   YP_T21 : TIMER[30] := ([0].PRE := 1000, [1].PRE := 10000000, [2].PRE := 10000000, [3].PRE := 3000, [3].ACC := 1845, [3].EN := 1, [3].TT := 1);
   YP_T4 : TIMER[16] := ([0].PRE := 3000, [0].ACC := 368, [0].EN := 1, [0].TT := 1, [1].PRE := 10000, [2].PRE := 10000, [2].ACC := 10001, [2].EN := 1, [2].DN := 1, [3].PRE := 60000, [3].ACC := 30907, [3].EN := 1, [3].TT := 1, [4].PRE := 5000, [4].ACC := 5000, [4].EN := 1, [4].DN := 1, [5].PRE := 5000, [6].PRE := 5000, [6].ACC := 5000, [6].EN := 1, [6].DN := 1, [7].PRE := 5000, [10].PRE := 1000);   // TIMER
        [4]   // YST1 HIGH LEVEL DE-B TIMER OFF =WET
        [5]   // YST1 HIGH LEVEL DE-B TIMER
   YP_TANK_NUMBER : ALIAS FOR YP_N10[11];
   YP_TIMER_SELECTED : ALIAS FOR YP_N55[41];   // Blunger Drain Timer Select
   YP_WATER_FILL_IDLE : ALIAS FOR YP_N40[2].0;   // BLUNGER WATER FILL IDLE
   YP_WATER_FILL_RUNNING : ALIAS FOR YP_N40[2].1;   // Blunger Water Feed Running
   YP_WD : PlantItem;   // WD
   YP_WD_RawOutput : ALIAS FOR RIO_Rack_3:3:O.Data.14;   // YP_WD
   YP_YST1_ALARM : ALIAS FOR YP_N10[1].0;
   YP_YST1_HIGH_MESSAGE : ALIAS FOR YP_B92[1].0;
   YP_YST1_HL : PlantItem;   // YST1_HL
   YP_YST1_HL_ALARM : ALIAS FOR YP_N7[38].0;
   YP_YST1_HL_FLAG : ALIAS FOR YP_N7[40].0;   // YST1 HIGH LEVEL FLAG ON=WET
   YP_YST1_HL_RawInput : ALIAS FOR RIO_Rack_3:1:I.Data.1;   // YP_YST1_HL
   YP_YST1_HL_TIMER : ALIAS FOR YP_T4[4];   // YST1 HIGH LEVEL DE-B TIMER OFF =WET
   YP_YST1_HL_TIMER2 : ALIAS FOR YP_T4[5];   // YST1 HIGH LEVEL DE-B TIMER
   YP_YST2_ALARM : ALIAS FOR YP_N10[1].1;
   YP_YST2_HIGH_LEVEL_FLAG : ALIAS FOR YP_N7[40].1;   // YST2 HIGH LEVEL FLAG ON=WET
   YP_YST2_HIGH_MESSAGE : ALIAS FOR YP_B92[1].1;
   YP_YST2_HL : PlantItem;   // YST2_HL
   YP_YST2_HL_ALARM : ALIAS FOR YP_N7[38].1;
   YP_YST2_HL_RawInput : ALIAS FOR RIO_Rack_3:1:I.Data.3;   // YP_YST2_HL
   YP_YST2_HL_TIMER : ALIAS FOR YP_T4[6];
   YP_YST2_HL_TIMER2 : ALIAS FOR YP_T4[7];
   YST_BL_PMP_ON : BOOL;   // Blunger Pump
   YST_CIP_Conns_Confirmed : BOOL := 1;
   YST_Confirm_CIP_connected : BOOL;
   YST_Confirm_Vent_connected : BOOL;
   YST_Vent_Connection_Confirmed : BOOL;
   YSVFilling_transaction_locked_timer : TIMER := (PRE := 10000);
   YSVFilling_transaction_log : DINT;
   YSVFilling_transaction_log_delay : DINT;
   YSVFilling_transaction_log_Done : DINT := -1;
   YSVFilling_transaction_log_timer : TIMER := (PRE := 10000);
END_VAR

PROGRAM _1Second   (* main routine OneSecond *)

ROUTINE OneSecond   (* ladder *)
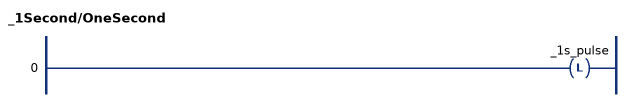
   0: OTL(_1s_pulse);
END_ROUTINE
END_PROGRAM

PROGRAM First_Task   (* main routine MainRoutine *)

ROUTINE MainRoutine   (* ladder *)
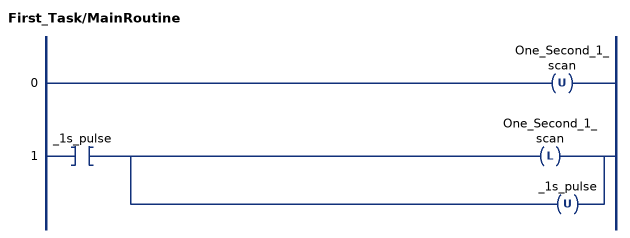
   0: OTU(One_Second_1_scan);
   1: XIC(_1s_pulse)[OTL(One_Second_1_scan) ,OTU(_1s_pulse) ];
END_ROUTINE
END_PROGRAM

PROGRAM FR_Common   (* main routine MainRoutine *)
VAR
   FR_FV31_AV08_O1 : ALIAS FOR RIO_Rack_2:12:I.Data.26;
   FR_FVS_P01_Cond_Met : BOOL;
END_VAR

ROUTINE A_FactoryTalk_Requirements   (* ladder *)
END_ROUTINE

ROUTINE Analog_scale_ftof   (* ladder *)
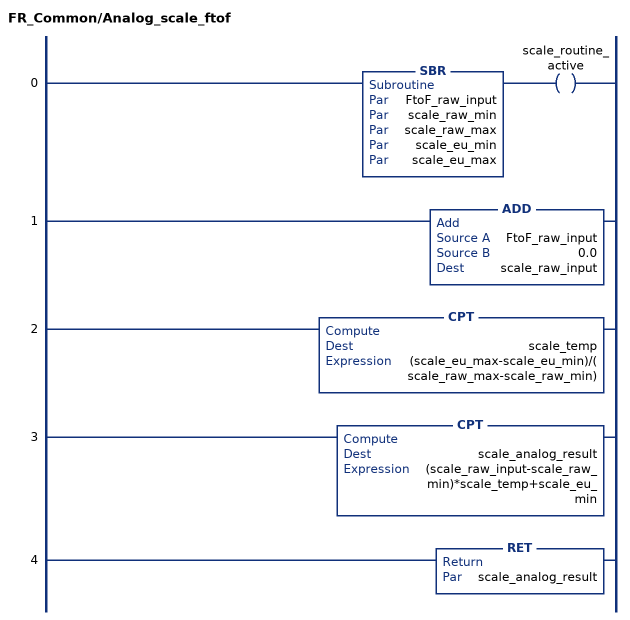
   0: SBR(FtoF_raw_input,scale_raw_min,scale_raw_max,scale_eu_min,scale_eu_max)OTE(scale_routine_active);
   1: ADD(FtoF_raw_input,0.0,scale_raw_input);
   2: CPT(scale_temp,(scale_eu_max-scale_eu_min)/(scale_raw_max-scale_raw_min));
   3: CPT(scale_analog_result,(scale_raw_input-scale_raw_min)*scale_temp+scale_eu_min);
   4: RET(scale_analog_result);
END_ROUTINE

ROUTINE Analog_Scale_FtoI   (* ladder *)
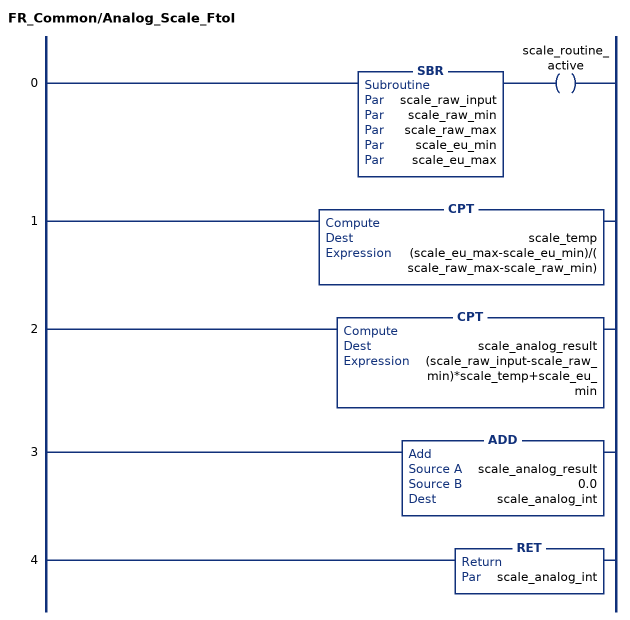
   0: SBR(scale_raw_input,scale_raw_min,scale_raw_max,scale_eu_min,scale_eu_max)OTE(scale_routine_active);
   1: CPT(scale_temp,(scale_eu_max-scale_eu_min)/(scale_raw_max-scale_raw_min));
   2: CPT(scale_analog_result,(scale_raw_input-scale_raw_min)*scale_temp+scale_eu_min);
   3: ADD(scale_analog_result,0.0,scale_analog_int);
   4: RET(scale_analog_int);
END_ROUTINE

ROUTINE Analog_Scale_ItoF   (* ladder *)
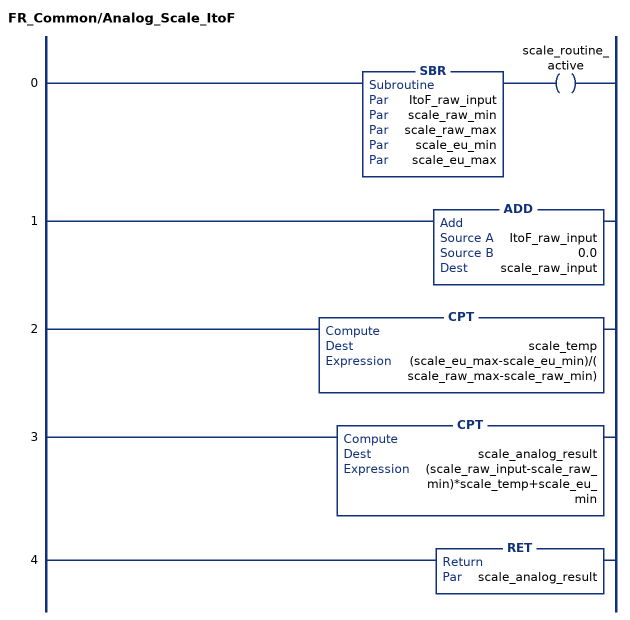
   0: SBR(ItoF_raw_input,scale_raw_min,scale_raw_max,scale_eu_min,scale_eu_max)OTE(scale_routine_active);
   1: ADD(ItoF_raw_input,0.0,scale_raw_input);
   2: CPT(scale_temp,(scale_eu_max-scale_eu_min)/(scale_raw_max-scale_raw_min));
   3: CPT(scale_analog_result,(scale_raw_input-scale_raw_min)*scale_temp+scale_eu_min);
   4: RET(scale_analog_result);
END_ROUTINE

ROUTINE Analog_Scale_ItoF_Int_Parms   (* ladder *)
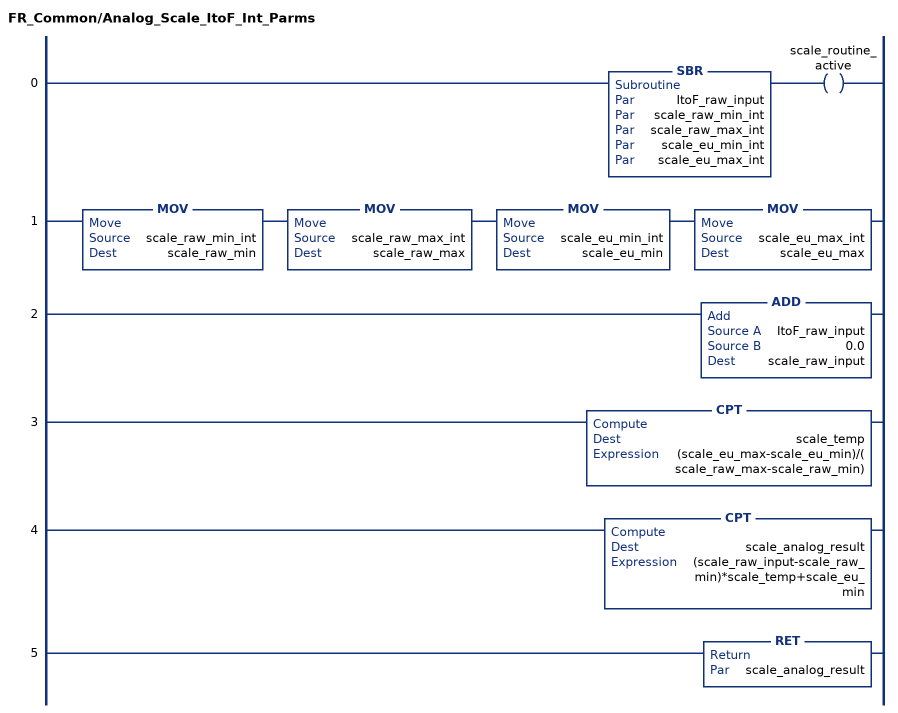
   0: SBR(ItoF_raw_input,scale_raw_min_int,scale_raw_max_int,scale_eu_min_int,scale_eu_max_int)OTE(scale_routine_active);
   1: MOV(scale_raw_min_int,scale_raw_min)MOV(scale_raw_max_int,scale_raw_max)MOV(scale_eu_min_int,scale_eu_min)MOV(scale_eu_max_int,scale_eu_max);
   2: ADD(ItoF_raw_input,0.0,scale_raw_input);
   3: CPT(scale_temp,(scale_eu_max-scale_eu_min)/(scale_raw_max-scale_raw_min));
   4: CPT(scale_analog_result,(scale_raw_input-scale_raw_min)*scale_temp+scale_eu_min);
   5: RET(scale_analog_result);
END_ROUTINE

ROUTINE FR_A_Alarms_From_PLC   (* ladder *)
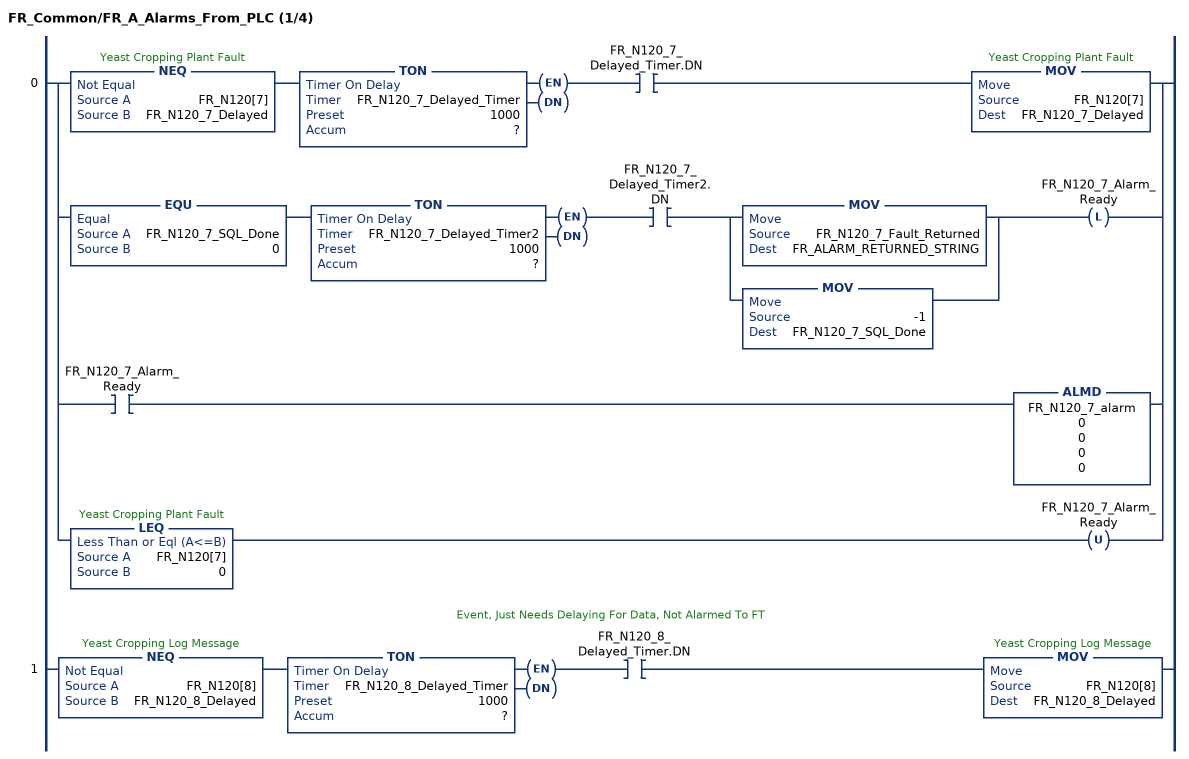
   0: [NEQ(FR_N120[7],FR_N120_7_Delayed) TON(FR_N120_7_Delayed_Timer,?,?) XIC(FR_N120_7_Delayed_Timer.DN) MOV(FR_N120[7],FR_N120_7_Delayed) ,EQU(FR_N120_7_SQL_Done,0) TON(FR_N120_7_Delayed_Timer2,?,?) XIC(FR_N120_7_Delayed_Timer2.DN) [MOV(FR_N120_7_Fault_Returned,FR_ALARM_RETURNED_STRING) ,MOV(-1,FR_N120_7_SQL_Done) ] OTL(FR_N120_7_Alarm_Ready) ,XIC(FR_N120_7_Alarm_Ready) ALMD(FR_N120_7_alarm,0,0,0,0) ,LEQ(FR_N120[7],0) OTU(FR_N120_7_Alarm_Ready) ];
   // Event, Just Needs Delaying For Data, Not Alarmed To FT
   1: NEQ(FR_N120[8],FR_N120_8_Delayed)TON(FR_N120_8_Delayed_Timer,?,?)XIC(FR_N120_8_Delayed_Timer.DN)MOV(FR_N120[8],FR_N120_8_Delayed);
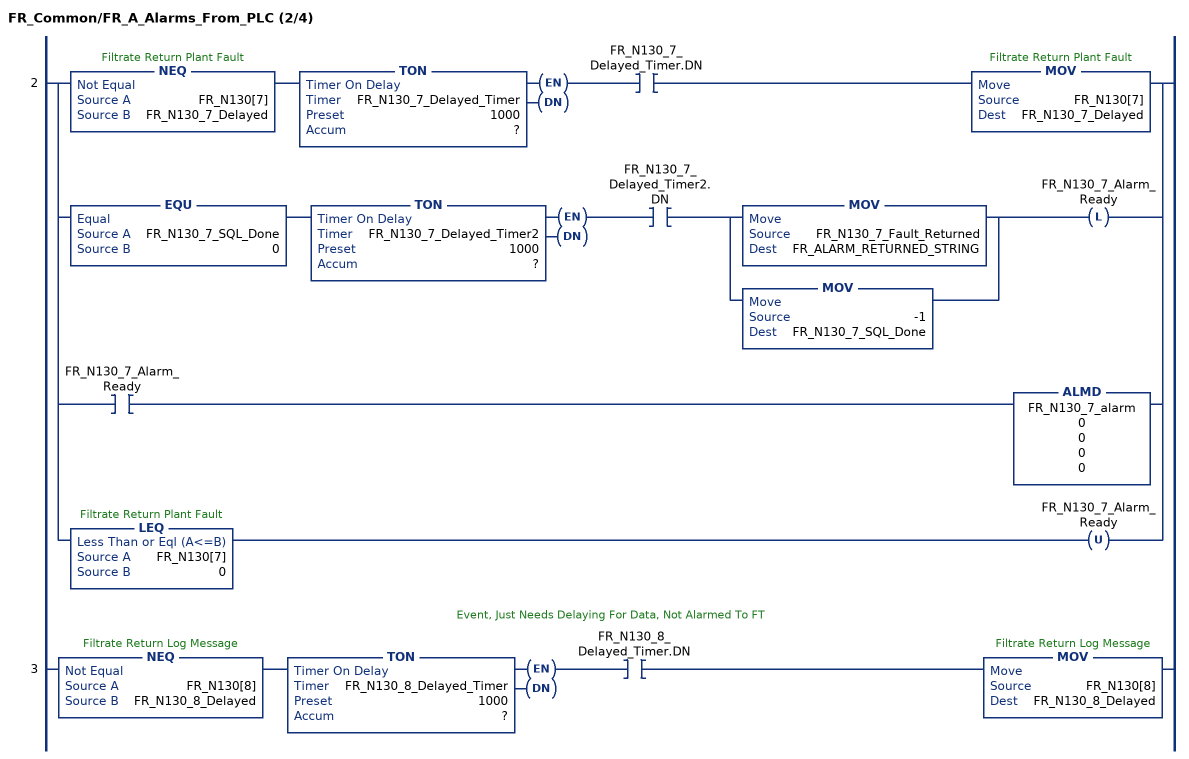
   2: [NEQ(FR_N130[7],FR_N130_7_Delayed) TON(FR_N130_7_Delayed_Timer,?,?) XIC(FR_N130_7_Delayed_Timer.DN) MOV(FR_N130[7],FR_N130_7_Delayed) ,EQU(FR_N130_7_SQL_Done,0) TON(FR_N130_7_Delayed_Timer2,?,?) XIC(FR_N130_7_Delayed_Timer2.DN) [MOV(FR_N130_7_Fault_Returned,FR_ALARM_RETURNED_STRING) ,MOV(-1,FR_N130_7_SQL_Done) ] OTL(FR_N130_7_Alarm_Ready) ,XIC(FR_N130_7_Alarm_Ready) ALMD(FR_N130_7_alarm,0,0,0,0) ,LEQ(FR_N130[7],0) OTU(FR_N130_7_Alarm_Ready) ];
   // Event, Just Needs Delaying For Data, Not Alarmed To FT
   3: NEQ(FR_N130[8],FR_N130_8_Delayed)TON(FR_N130_8_Delayed_Timer,?,?)XIC(FR_N130_8_Delayed_Timer.DN)MOV(FR_N130[8],FR_N130_8_Delayed);
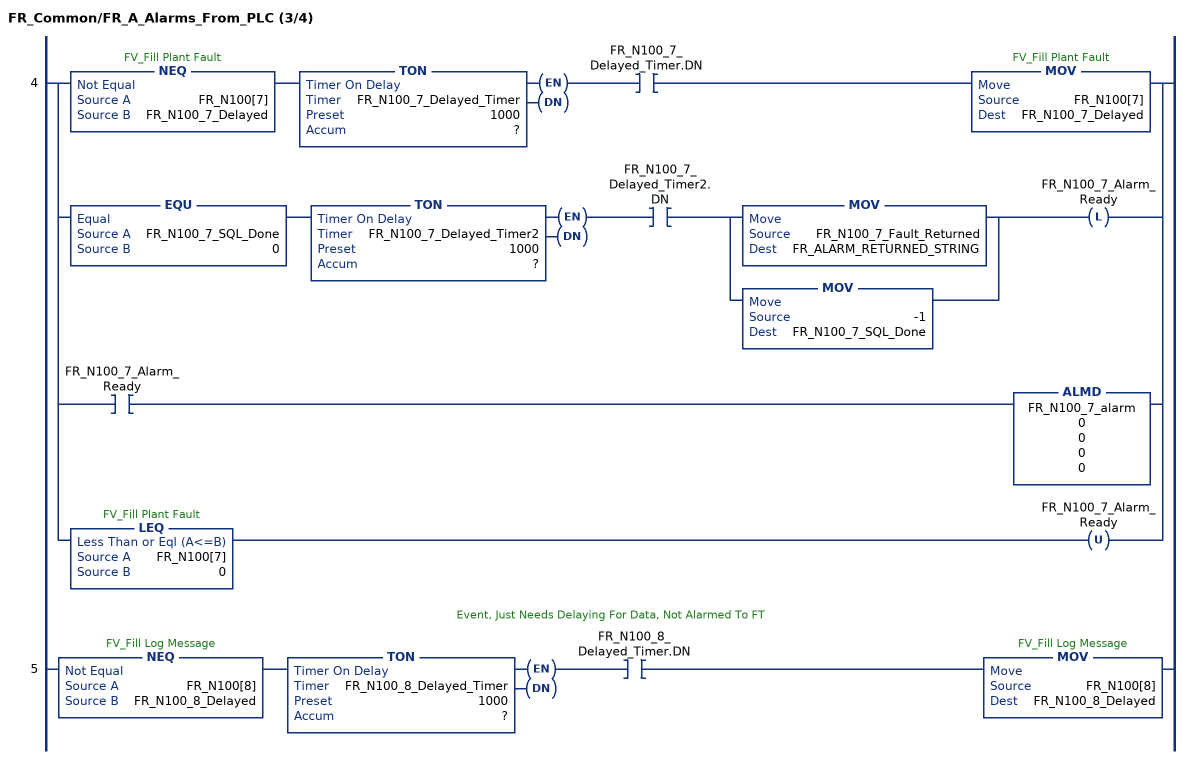
   4: [NEQ(FR_N100[7],FR_N100_7_Delayed) TON(FR_N100_7_Delayed_Timer,?,?) XIC(FR_N100_7_Delayed_Timer.DN) MOV(FR_N100[7],FR_N100_7_Delayed) ,EQU(FR_N100_7_SQL_Done,0) TON(FR_N100_7_Delayed_Timer2,?,?) XIC(FR_N100_7_Delayed_Timer2.DN) [MOV(FR_N100_7_Fault_Returned,FR_ALARM_RETURNED_STRING) ,MOV(-1,FR_N100_7_SQL_Done) ] OTL(FR_N100_7_Alarm_Ready) ,XIC(FR_N100_7_Alarm_Ready) ALMD(FR_N100_7_alarm,0,0,0,0) ,LEQ(FR_N100[7],0) OTU(FR_N100_7_Alarm_Ready) ];
   // Event, Just Needs Delaying For Data, Not Alarmed To FT
   5: NEQ(FR_N100[8],FR_N100_8_Delayed)TON(FR_N100_8_Delayed_Timer,?,?)XIC(FR_N100_8_Delayed_Timer.DN)MOV(FR_N100[8],FR_N100_8_Delayed);
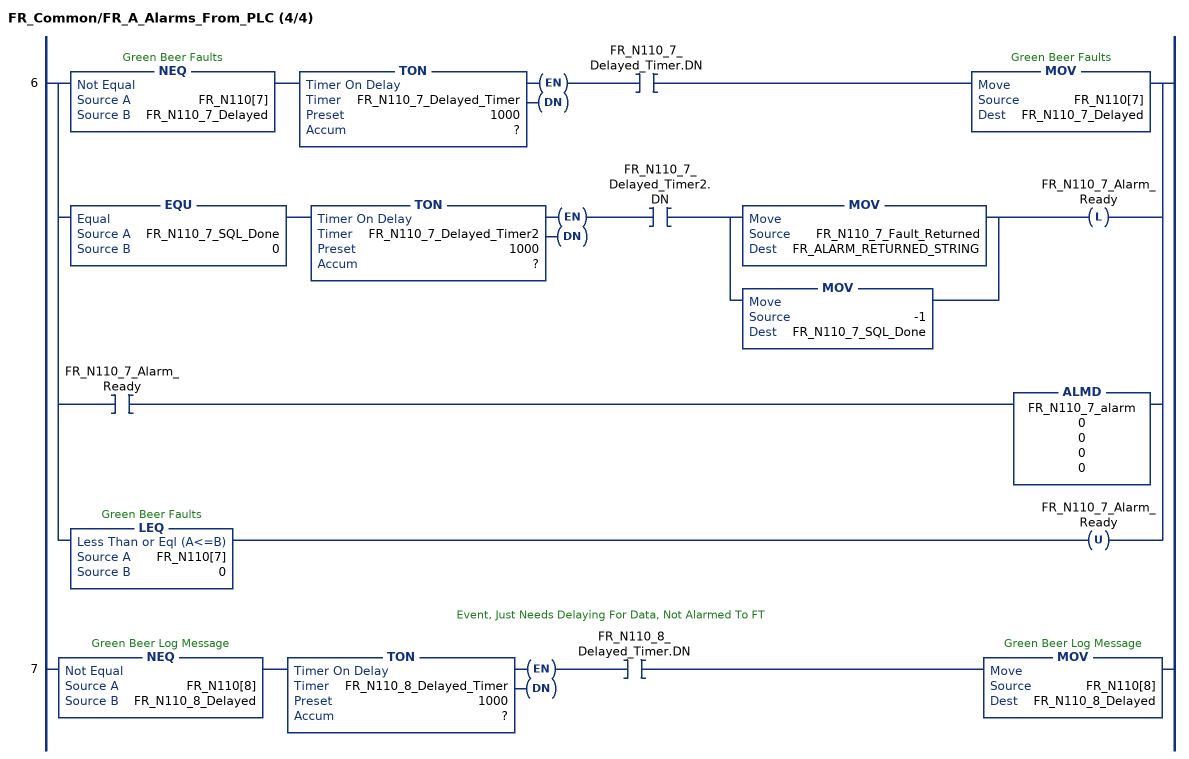
   6: [NEQ(FR_N110[7],FR_N110_7_Delayed) TON(FR_N110_7_Delayed_Timer,?,?) XIC(FR_N110_7_Delayed_Timer.DN) MOV(FR_N110[7],FR_N110_7_Delayed) ,EQU(FR_N110_7_SQL_Done,0) TON(FR_N110_7_Delayed_Timer2,?,?) XIC(FR_N110_7_Delayed_Timer2.DN) [MOV(FR_N110_7_Fault_Returned,FR_ALARM_RETURNED_STRING) ,MOV(-1,FR_N110_7_SQL_Done) ] OTL(FR_N110_7_Alarm_Ready) ,XIC(FR_N110_7_Alarm_Ready) ALMD(FR_N110_7_alarm,0,0,0,0) ,LEQ(FR_N110[7],0) OTU(FR_N110_7_Alarm_Ready) ];
   // Event, Just Needs Delaying For Data, Not Alarmed To FT
   7: NEQ(FR_N110[8],FR_N110_8_Delayed)TON(FR_N110_8_Delayed_Timer,?,?)XIC(FR_N110_8_Delayed_Timer.DN)MOV(FR_N110[8],FR_N110_8_Delayed);
END_ROUTINE

ROUTINE FR_A_Events_From_Scada   (* ladder *)
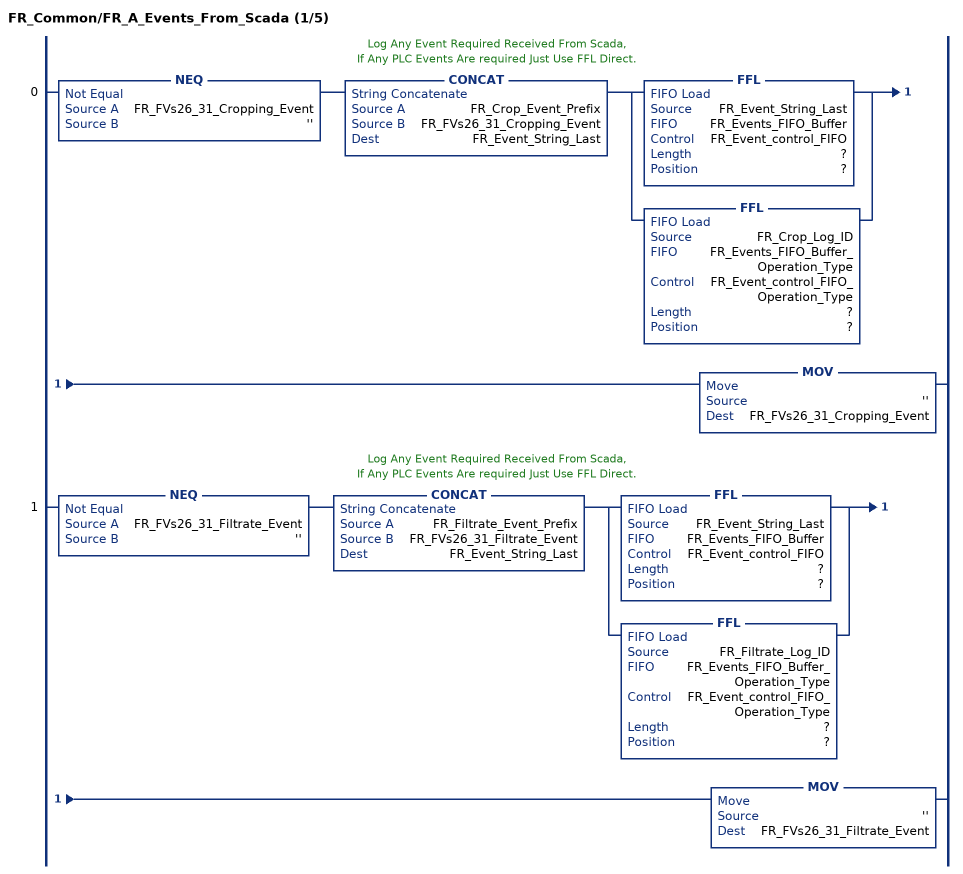
   // Log Any Event Required Received From Scada,
   // If Any PLC Events Are required Just Use FFL Direct.
   0: NEQ(FR_FVs26_31_Cropping_Event,'')CONCAT(FR_Crop_Event_Prefix,FR_FVs26_31_Cropping_Event,FR_Event_String_Last)[FFL(FR_Event_String_Last,FR_Events_FIFO_Buffer,FR_Event_control_FIFO,?,?) ,FFL(FR_Crop_Log_ID,FR_Events_FIFO_Buffer_Operation_Type,FR_Event_control_FIFO_Operation_Type,?,?) ]MOV('',FR_FVs26_31_Cropping_Event);
   // Log Any Event Required Received From Scada,
   // If Any PLC Events Are required Just Use FFL Direct.
   1: NEQ(FR_FVs26_31_Filtrate_Event,'')CONCAT(FR_Filtrate_Event_Prefix,FR_FVs26_31_Filtrate_Event,FR_Event_String_Last)[FFL(FR_Event_String_Last,FR_Events_FIFO_Buffer,FR_Event_control_FIFO,?,?) ,FFL(FR_Filtrate_Log_ID,FR_Events_FIFO_Buffer_Operation_Type,FR_Event_control_FIFO_Operation_Type,?,?) ]MOV('',FR_FVs26_31_Filtrate_Event);
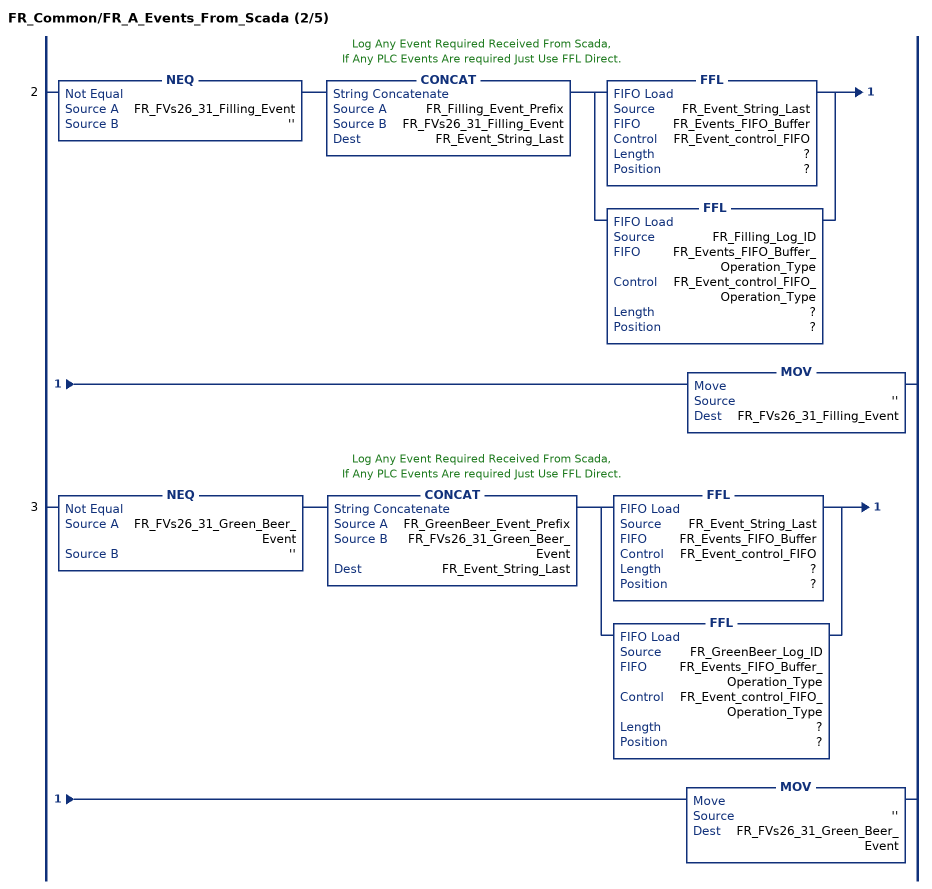
   // Log Any Event Required Received From Scada,
   // If Any PLC Events Are required Just Use FFL Direct.
   2: NEQ(FR_FVs26_31_Filling_Event,'')CONCAT(FR_Filling_Event_Prefix,FR_FVs26_31_Filling_Event,FR_Event_String_Last)[FFL(FR_Event_String_Last,FR_Events_FIFO_Buffer,FR_Event_control_FIFO,?,?) ,FFL(FR_Filling_Log_ID,FR_Events_FIFO_Buffer_Operation_Type,FR_Event_control_FIFO_Operation_Type,?,?) ]MOV('',FR_FVs26_31_Filling_Event);
   // Log Any Event Required Received From Scada,
   // If Any PLC Events Are required Just Use FFL Direct.
   3: NEQ(FR_FVs26_31_Green_Beer_Event,'')CONCAT(FR_GreenBeer_Event_Prefix,FR_FVs26_31_Green_Beer_Event,FR_Event_String_Last)[FFL(FR_Event_String_Last,FR_Events_FIFO_Buffer,FR_Event_control_FIFO,?,?) ,FFL(FR_GreenBeer_Log_ID,FR_Events_FIFO_Buffer_Operation_Type,FR_Event_control_FIFO_Operation_Type,?,?) ]MOV('',FR_FVs26_31_Green_Beer_Event);
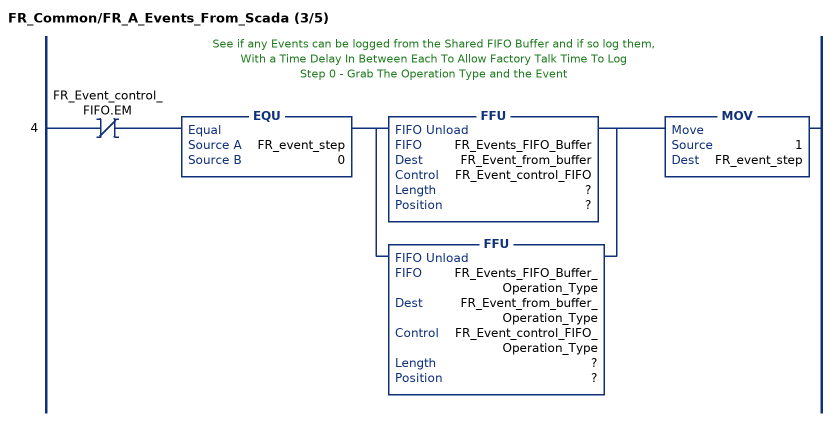
   // See if any Events can be logged from the Shared FIFO Buffer and if so log them,
   // With a Time Delay In Between Each To Allow Factory Talk Time To Log
   // Step 0 - Grab The Operation Type and the Event
   4: XIO(FR_Event_control_FIFO.EM)EQU(FR_event_step,0)[FFU(FR_Events_FIFO_Buffer,FR_Event_from_buffer,FR_Event_control_FIFO,?,?) ,FFU(FR_Events_FIFO_Buffer_Operation_Type,FR_Event_from_buffer_Operation_Type,FR_Event_control_FIFO_Operation_Type,?,?) ]MOV(1,FR_event_step);
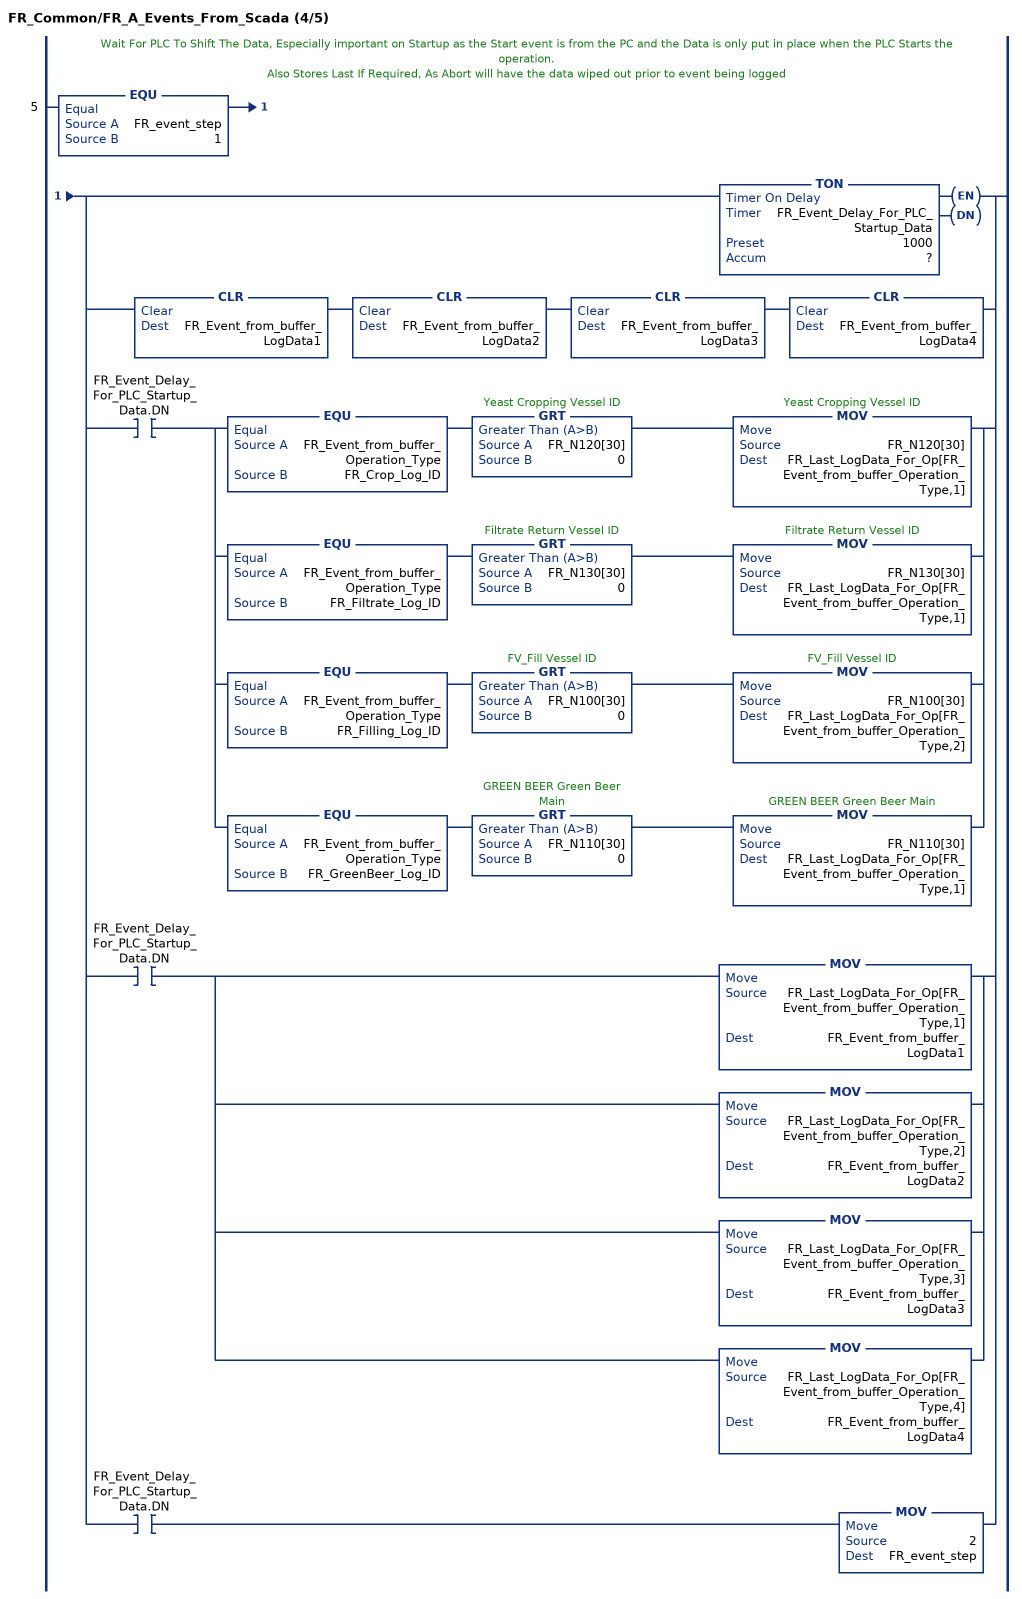
   // Wait For PLC To Shift The Data, Especially important on Startup as the Start event is from the PC and the Data is only put in place when the PLC Starts the operation.
   // Also Stores Last If Required, As Abort will have the data wiped out prior to event being logged
   5: EQU(FR_event_step,1)[TON(FR_Event_Delay_For_PLC_Startup_Data,?,?) ,CLR(FR_Event_from_buffer_LogData1) CLR(FR_Event_from_buffer_LogData2) CLR(FR_Event_from_buffer_LogData3) CLR(FR_Event_from_buffer_LogData4) ,XIC(FR_Event_Delay_For_PLC_Startup_Data.DN) [EQU(FR_Event_from_buffer_Operation_Type,FR_Crop_Log_ID) GRT(FR_N120[30],0) MOV(FR_N120[30],FR_Last_LogData_For_Op[FR_Event_from_buffer_Operation_Type,1]) ,EQU(FR_Event_from_buffer_Operation_Type,FR_Filtrate_Log_ID) GRT(FR_N130[30],0) MOV(FR_N130[30],FR_Last_LogData_For_Op[FR_Event_from_buffer_Operation_Type,1]) ,EQU(FR_Event_from_buffer_Operation_Type,FR_Filling_Log_ID) GRT(FR_N100[30],0) MOV(FR_N100[30],FR_Last_LogData_For_Op[FR_Event_from_buffer_Operation_Type,2]) ,EQU(FR_Event_from_buffer_Operation_Type,FR_GreenBeer_Log_ID) GRT(FR_N110[30],0) MOV(FR_N110[30],FR_Last_LogData_For_Op[FR_Event_from_buffer_Operation_Type,1]) ] ,XIC(FR_Event_Delay_For_PLC_Startup_Data.DN) [MOV(FR_Last_LogData_For_Op[FR_Event_from_buffer_Operation_Type,1],FR_Event_from_buffer_LogData1) ,MOV(FR_Last_LogData_For_Op[FR_Event_from_buffer_Operation_Type,2],FR_Event_from_buffer_LogData2) ,MOV(FR_Last_LogData_For_Op[FR_Event_from_buffer_Operation_Type,3],FR_Event_from_buffer_LogData3) ,MOV(FR_Last_LogData_For_Op[FR_Event_from_buffer_Operation_Type,4],FR_Event_from_buffer_LogData4) ] ,XIC(FR_Event_Delay_For_PLC_Startup_Data.DN) MOV(2,FR_event_step) ];
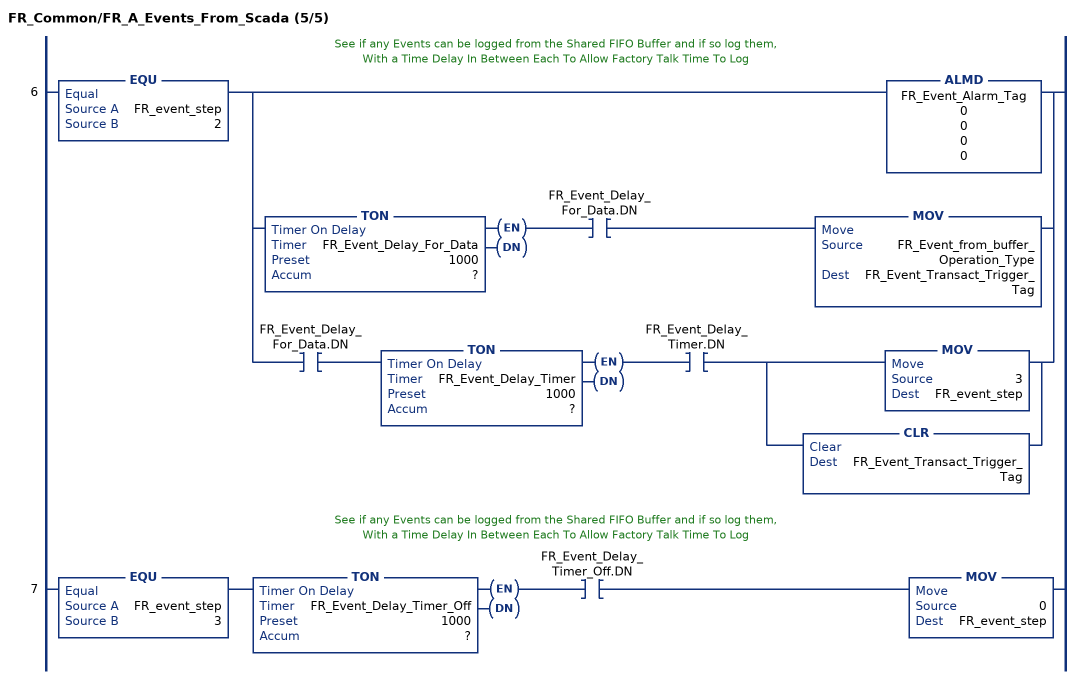
   // See if any Events can be logged from the Shared FIFO Buffer and if so log them,
   // With a Time Delay In Between Each To Allow Factory Talk Time To Log
   6: EQU(FR_event_step,2)[ALMD(FR_Event_Alarm_Tag,0,0,0,0) ,TON(FR_Event_Delay_For_Data,?,?) XIC(FR_Event_Delay_For_Data.DN) MOV(FR_Event_from_buffer_Operation_Type,FR_Event_Transact_Trigger_Tag) ,XIC(FR_Event_Delay_For_Data.DN) TON(FR_Event_Delay_Timer,?,?) XIC(FR_Event_Delay_Timer.DN) [MOV(3,FR_event_step) ,CLR(FR_Event_Transact_Trigger_Tag) ] ];
   // See if any Events can be logged from the Shared FIFO Buffer and if so log them,
   // With a Time Delay In Between Each To Allow Factory Talk Time To Log
   7: EQU(FR_event_step,3)TON(FR_Event_Delay_Timer_Off,?,?)XIC(FR_Event_Delay_Timer_Off.DN)MOV(0,FR_event_step);
END_ROUTINE

ROUTINE FR_A_Events_From_Scada_IDs   (* ladder *)
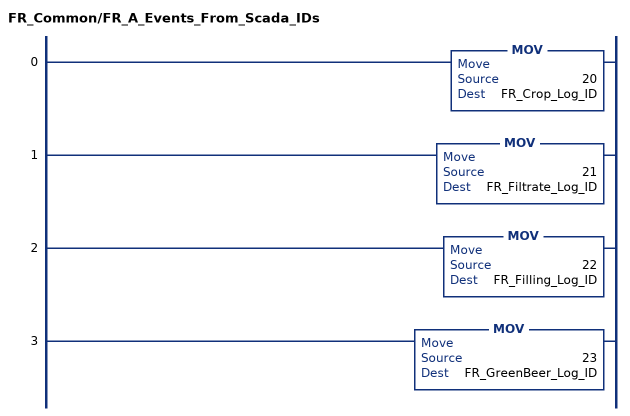
   0: MOV(20,FR_Crop_Log_ID);
   1: MOV(21,FR_Filtrate_Log_ID);
   2: MOV(22,FR_Filling_Log_ID);
   3: MOV(23,FR_GreenBeer_Log_ID);
END_ROUTINE

ROUTINE FR_A_Warnings_From_PLC   (* ladder *)
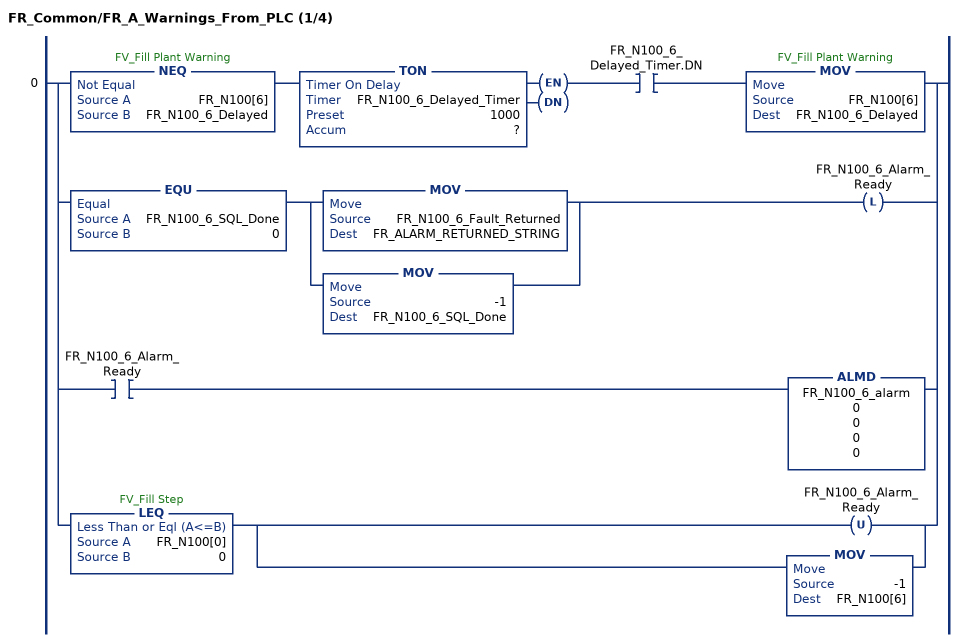
   0: [NEQ(FR_N100[6],FR_N100_6_Delayed) TON(FR_N100_6_Delayed_Timer,?,?) XIC(FR_N100_6_Delayed_Timer.DN) MOV(FR_N100[6],FR_N100_6_Delayed) ,EQU(FR_N100_6_SQL_Done,0) [MOV(FR_N100_6_Fault_Returned,FR_ALARM_RETURNED_STRING) ,MOV(-1,FR_N100_6_SQL_Done) ] OTL(FR_N100_6_Alarm_Ready) ,XIC(FR_N100_6_Alarm_Ready) ALMD(FR_N100_6_alarm,0,0,0,0) ,LEQ(FR_N100[0],0) [OTU(FR_N100_6_Alarm_Ready) ,MOV(-1,FR_N100[6]) ] ];
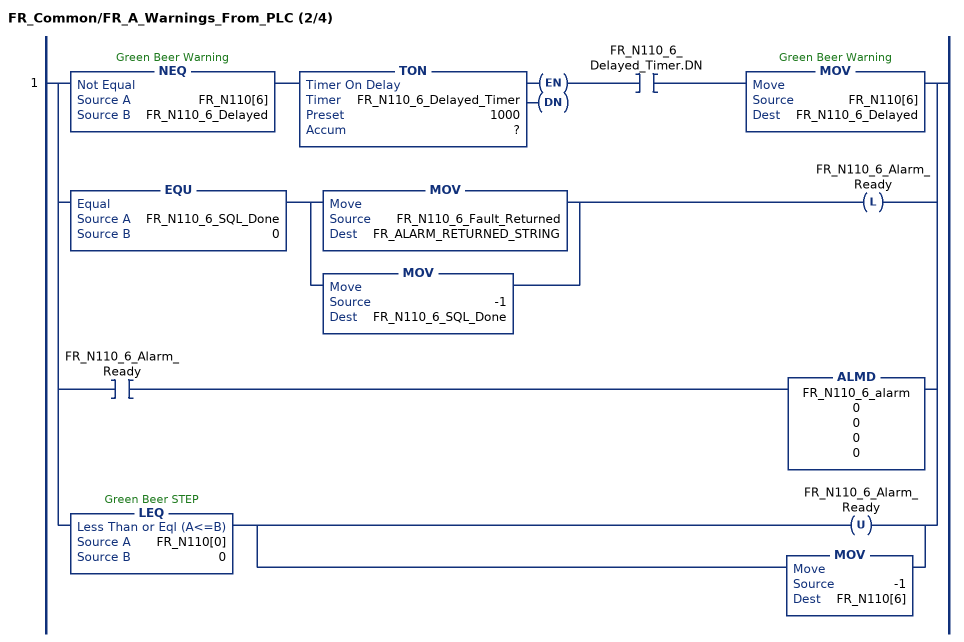
   1: [NEQ(FR_N110[6],FR_N110_6_Delayed) TON(FR_N110_6_Delayed_Timer,?,?) XIC(FR_N110_6_Delayed_Timer.DN) MOV(FR_N110[6],FR_N110_6_Delayed) ,EQU(FR_N110_6_SQL_Done,0) [MOV(FR_N110_6_Fault_Returned,FR_ALARM_RETURNED_STRING) ,MOV(-1,FR_N110_6_SQL_Done) ] OTL(FR_N110_6_Alarm_Ready) ,XIC(FR_N110_6_Alarm_Ready) ALMD(FR_N110_6_alarm,0,0,0,0) ,LEQ(FR_N110[0],0) [OTU(FR_N110_6_Alarm_Ready) ,MOV(-1,FR_N110[6]) ] ];
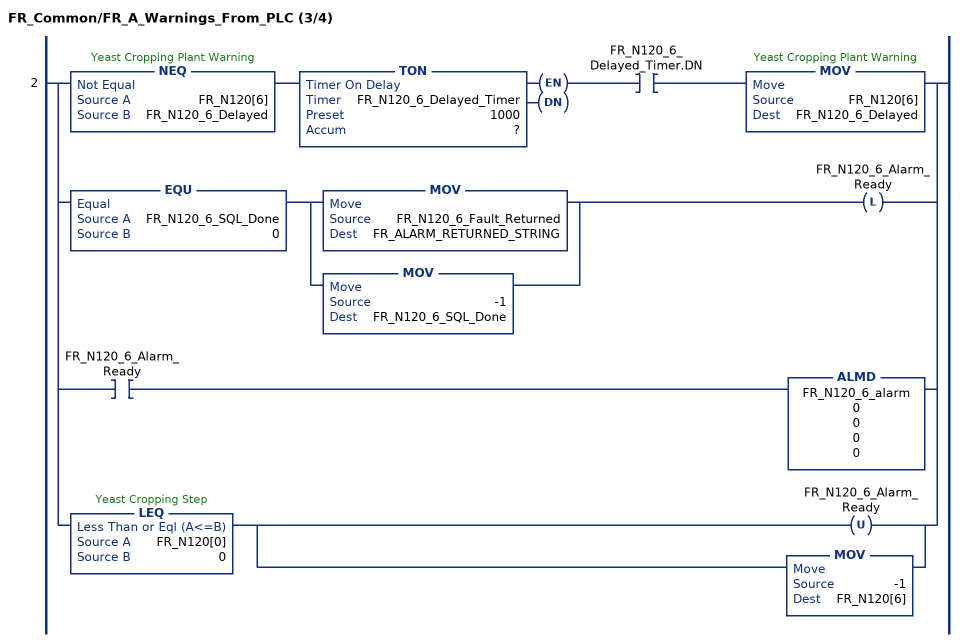
   2: [NEQ(FR_N120[6],FR_N120_6_Delayed) TON(FR_N120_6_Delayed_Timer,?,?) XIC(FR_N120_6_Delayed_Timer.DN) MOV(FR_N120[6],FR_N120_6_Delayed) ,EQU(FR_N120_6_SQL_Done,0) [MOV(FR_N120_6_Fault_Returned,FR_ALARM_RETURNED_STRING) ,MOV(-1,FR_N120_6_SQL_Done) ] OTL(FR_N120_6_Alarm_Ready) ,XIC(FR_N120_6_Alarm_Ready) ALMD(FR_N120_6_alarm,0,0,0,0) ,LEQ(FR_N120[0],0) [OTU(FR_N120_6_Alarm_Ready) ,MOV(-1,FR_N120[6]) ] ];
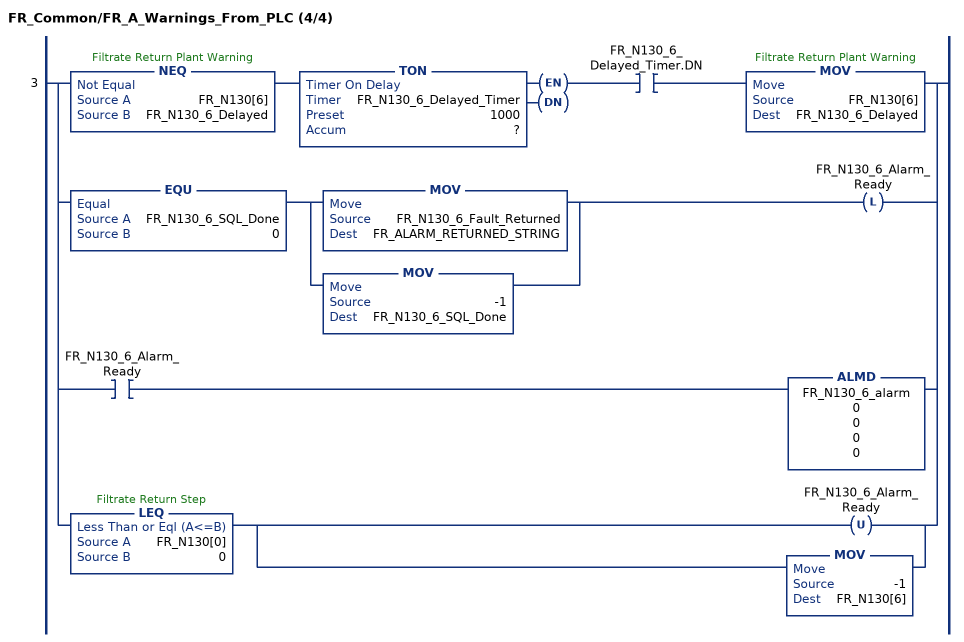
   3: [NEQ(FR_N130[6],FR_N130_6_Delayed) TON(FR_N130_6_Delayed_Timer,?,?) XIC(FR_N130_6_Delayed_Timer.DN) MOV(FR_N130[6],FR_N130_6_Delayed) ,EQU(FR_N130_6_SQL_Done,0) [MOV(FR_N130_6_Fault_Returned,FR_ALARM_RETURNED_STRING) ,MOV(-1,FR_N130_6_SQL_Done) ] OTL(FR_N130_6_Alarm_Ready) ,XIC(FR_N130_6_Alarm_Ready) ALMD(FR_N130_6_alarm,0,0,0,0) ,LEQ(FR_N130[0],0) [OTU(FR_N130_6_Alarm_Ready) ,MOV(-1,FR_N130[6]) ] ];
END_ROUTINE
